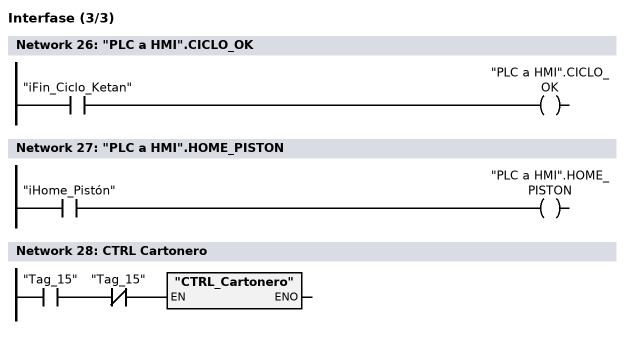
   RUNG wire#powerrail
      Contact( "iFin_Ciclo_Ketan" )
      Coil( "PLC a HMI".CICLO_OK )
   END_RUNG
   // the same network as SCL:
   "PLC a HMI".CICLO_OK := "iFin_Ciclo_Ketan";
END_REGION

REGION Network 27: "PLC a HMI".HOME_PISTON
   RUNG wire#powerrail
      Contact( "iHome_Pistón" )
      Coil( "PLC a HMI".HOME_PISTON )
   END_RUNG
   // the same network as SCL:
   "PLC a HMI".HOME_PISTON := "iHome_Pistón";
END_REGION

REGION Network 28: CTRL Cartonero
   RUNG wire#powerrail
      Contact( "Tag_15" )
      I_Contact( "Tag_15" )
      "CTRL_Cartonero"()
   END_RUNG
   // the same network as SCL:
   IF "Tag_15" AND NOT "Tag_15" THEN "CTRL_Cartonero"(); END_IF;
END_REGION
END_FUNCTION

FUNCTION "Conteo_AUTO" : Void   // FC26, STL
{ S7_Optimized_Access := 'FALSE' }
VERSION : 0.1
BEGIN

REGION Network 1: "Proceso CargaPallet".Capa_Actual
   // Con el fp del empujador adelante de todo, actualiza la "Capa_Actual" del grupo "CargaPalet"
         A     "flanco".piSnsEmpj_Ade_Par;
         JCN   NoCapa;
         L     "Proceso Empujador".Capa_Actual;
         T     "Proceso CargaPallet".Capa_Actual;
   NoCapa:NOP   0;
END_REGION

REGION Network 2
         L     "DB_Receta_Actual".Nro_Capas_Pallet;
         L     "Proceso Empujador".Capa_Actual;
         >I;
         =     #Habil_Inc;
         ==I;
         =     #Fin_Pallet;
         SET;
         A     #Habil_Inc;
         A     "flanco".piSnsEmpj_Ade_Par;
         JCN   noInc;
         L     "Proceso Empujador".Capa_Actual;
         INC   1;
         T     "Proceso Empujador".Capa_Actual;
   noInc:NOP   0;
         SET;
         A     #Fin_Pallet;
         A     "flanco".piSnsEmpj_Ade_Par;

         JCN   noFin;
         SET;
         S     "Última_Capa";
         L     1;
         T     "Proceso Empujador".Capa_Actual;
         L     "Proceso Empujador".Cant_Pallets;
         INC   1;
         T     "Proceso Empujador".Cant_Pallets;
   noFin:NOP   0;

         A     "flanco".nPALLET_NO_FUERA_ASCENSOR;
         JCN   noWRPall;
         L     "Proceso Empujador".Cant_Pallets;
         T     "Proceso CargaPallet".Cant_Pallets;
   noWRPall:NOP   0;


   //////////////////////////////
   //      O     "Ascensor_Zona_Superior"//
   //U     "flanco".nPALLET_NO_FUERA_ASCENSOR
   //     R     "Última_Capa"
END_REGION
END_FUNCTION

FUNCTION "Filtros_Señales" : Void   // FC27, LAD
{ S7_Optimized_Access := 'FALSE' }
VERSION : 0.1
BEGIN

REGION Network 1: Sensor Contador de embalaje 1
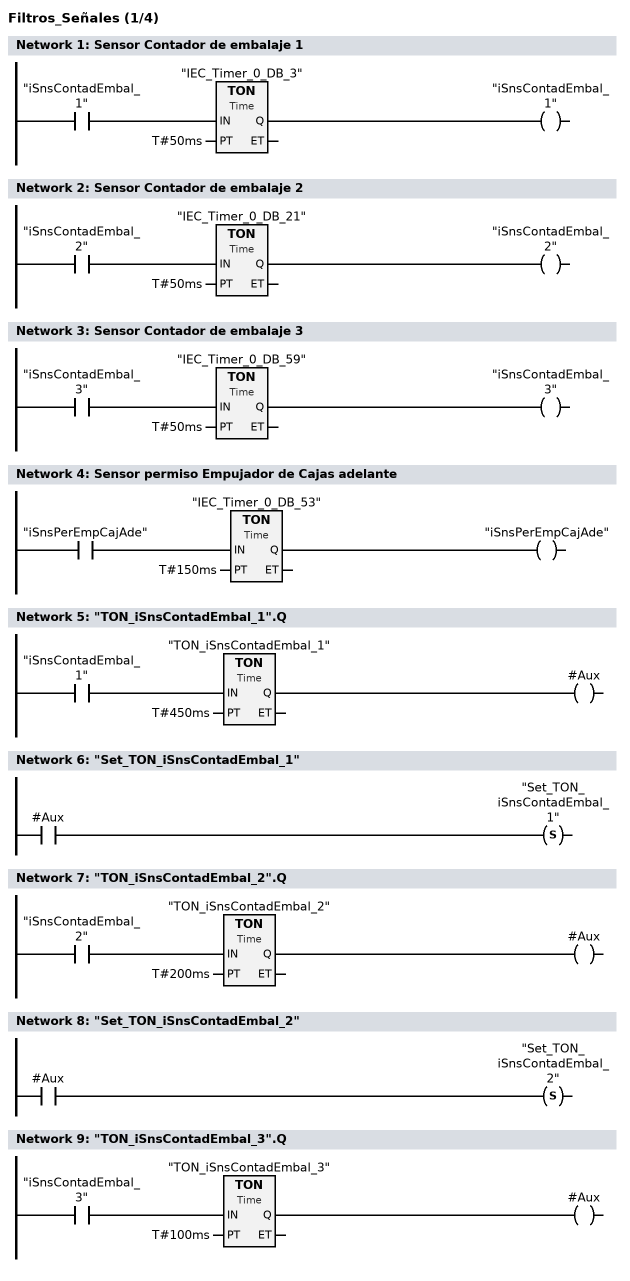
   "IEC_Timer_0_DB_3".TON(IN := "iSnsContadEmbal_1", PT := T#50ms);
   "iSnsContadEmbal_1" := "IEC_Timer_0_DB_3".Q;
END_REGION

REGION Network 2: Sensor Contador de embalaje 2
   "IEC_Timer_0_DB_21".TON(IN := "iSnsContadEmbal_2", PT := T#50ms);
   "iSnsContadEmbal_2" := "IEC_Timer_0_DB_21".Q;
END_REGION

REGION Network 3: Sensor Contador de embalaje 3
   "IEC_Timer_0_DB_59".TON(IN := "iSnsContadEmbal_3", PT := T#50ms);
   "iSnsContadEmbal_3" := "IEC_Timer_0_DB_59".Q;
END_REGION

REGION Network 4: Sensor permiso Empujador de Cajas adelante
   "IEC_Timer_0_DB_53".TON(IN := "iSnsPerEmpCajAde", PT := T#150ms);
   "iSnsPerEmpCajAde" := "IEC_Timer_0_DB_53".Q;
END_REGION

REGION Network 5: "TON_iSnsContadEmbal_1".Q
   "TON_iSnsContadEmbal_1".TON(IN := "iSnsContadEmbal_1", PT := T#450ms);
   #Aux := "TON_iSnsContadEmbal_1".Q;
END_REGION

REGION Network 6: "Set_TON_iSnsContadEmbal_1"
   RUNG wire#powerrail
      Contact( #Aux )
      S_Coil( "Set_TON_iSnsContadEmbal_1" )
   END_RUNG
   // the same network as SCL:
   IF #Aux THEN "Set_TON_iSnsContadEmbal_1" := TRUE; END_IF;
END_REGION

REGION Network 7: "TON_iSnsContadEmbal_2".Q
   "TON_iSnsContadEmbal_2".TON(IN := "iSnsContadEmbal_2", PT := T#200ms);
   #Aux := "TON_iSnsContadEmbal_2".Q;
END_REGION

REGION Network 8: "Set_TON_iSnsContadEmbal_2"
   RUNG wire#powerrail
      Contact( #Aux )
      S_Coil( "Set_TON_iSnsContadEmbal_2" )
   END_RUNG
   // the same network as SCL:
   IF #Aux THEN "Set_TON_iSnsContadEmbal_2" := TRUE; END_IF;
END_REGION

REGION Network 9: "TON_iSnsContadEmbal_3".Q
   "TON_iSnsContadEmbal_3".TON(IN := "iSnsContadEmbal_3", PT := T#100ms);
   #Aux := "TON_iSnsContadEmbal_3".Q;
END_REGION

REGION Network 10: "Set_TON_iSnsContadEmbal_3"
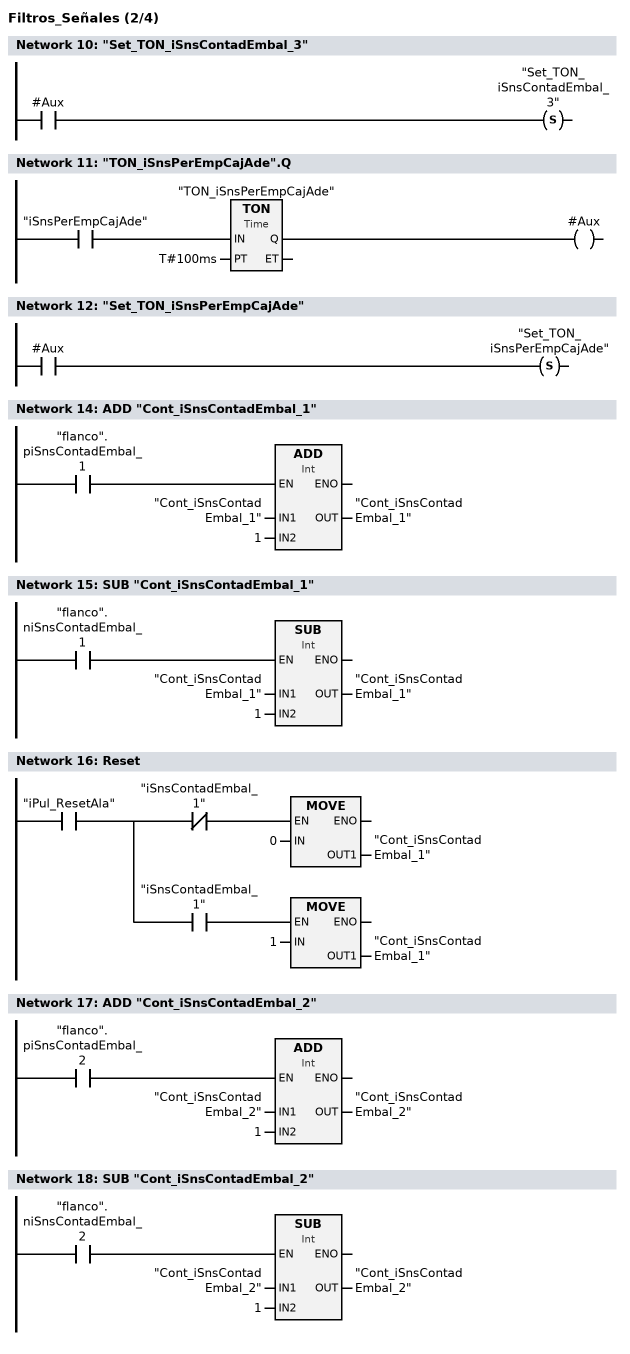
   RUNG wire#powerrail
      Contact( #Aux )
      S_Coil( "Set_TON_iSnsContadEmbal_3" )
   END_RUNG
   // the same network as SCL:
   IF #Aux THEN "Set_TON_iSnsContadEmbal_3" := TRUE; END_IF;
END_REGION

REGION Network 11: "TON_iSnsPerEmpCajAde".Q
   "TON_iSnsPerEmpCajAde".TON(IN := "iSnsPerEmpCajAde", PT := T#100ms);
   #Aux := "TON_iSnsPerEmpCajAde".Q;
END_REGION

REGION Network 12: "Set_TON_iSnsPerEmpCajAde"
   RUNG wire#powerrail
      Contact( #Aux )
      S_Coil( "Set_TON_iSnsPerEmpCajAde" )
   END_RUNG
   // the same network as SCL:
   IF #Aux THEN "Set_TON_iSnsPerEmpCajAde" := TRUE; END_IF;
END_REGION

REGION Network 13: ------------------------------------------ Control de flancos -------------------------------------------------
END_REGION

REGION Network 14: ADD "Cont_iSnsContadEmbal_1"
   RUNG wire#powerrail
      Contact( "flanco".piSnsContadEmbal_1 )
      { S7_Templates := "SrcType := Int"; S7_GenerateENO := "TRUE" } Add(in1 := "Cont_iSnsContadEmbal_1", in2 := 1, out => "Cont_iSnsContadEmbal_1")
   END_RUNG
   // the same network as SCL:
   IF "flanco".piSnsContadEmbal_1 THEN "Cont_iSnsContadEmbal_1" := "Cont_iSnsContadEmbal_1" + 1; END_IF;
END_REGION

REGION Network 15: SUB "Cont_iSnsContadEmbal_1"
   RUNG wire#powerrail
      Contact( "flanco".niSnsContadEmbal_1 )
      { S7_Templates := "SrcType := Int"; S7_GenerateENO := "TRUE" } Sub(in1 := "Cont_iSnsContadEmbal_1", in2 := 1, out => "Cont_iSnsContadEmbal_1")
   END_RUNG
   // the same network as SCL:
   IF "flanco".niSnsContadEmbal_1 THEN "Cont_iSnsContadEmbal_1" := "Cont_iSnsContadEmbal_1" - 1; END_IF;
END_REGION

REGION Network 16: Reset
   RUNG wire#powerrail
      Contact( "iPul_ResetAla" )
      wire#w1
      I_Contact( "iSnsContadEmbal_1" )
      { S7_GenerateENO := "TRUE" } Move(in := 0, out1 => "Cont_iSnsContadEmbal_1")
   END_RUNG
   RUNG wire#w1
      Contact( "iSnsContadEmbal_1" )
      { S7_GenerateENO := "TRUE" } Move(in := 1, out1 => "Cont_iSnsContadEmbal_1")
   END_RUNG
   // the same network as SCL:
   IF "iPul_ResetAla" AND NOT "iSnsContadEmbal_1" THEN "Cont_iSnsContadEmbal_1" := 0; END_IF;
   IF "iPul_ResetAla" AND "iSnsContadEmbal_1" THEN "Cont_iSnsContadEmbal_1" := 1; END_IF;
END_REGION

REGION Network 17: ADD "Cont_iSnsContadEmbal_2"
   RUNG wire#powerrail
      Contact( "flanco".piSnsContadEmbal_2 )
      { S7_Templates := "SrcType := Int"; S7_GenerateENO := "TRUE" } Add(in1 := "Cont_iSnsContadEmbal_2", in2 := 1, out => "Cont_iSnsContadEmbal_2")
   END_RUNG
   // the same network as SCL:
   IF "flanco".piSnsContadEmbal_2 THEN "Cont_iSnsContadEmbal_2" := "Cont_iSnsContadEmbal_2" + 1; END_IF;
END_REGION

REGION Network 18: SUB "Cont_iSnsContadEmbal_2"
   RUNG wire#powerrail
      Contact( "flanco".niSnsContadEmbal_2 )
      { S7_Templates := "SrcType := Int"; S7_GenerateENO := "TRUE" } Sub(in1 := "Cont_iSnsContadEmbal_2", in2 := 1, out => "Cont_iSnsContadEmbal_2")
   END_RUNG
   // the same network as SCL:
   IF "flanco".niSnsContadEmbal_2 THEN "Cont_iSnsContadEmbal_2" := "Cont_iSnsContadEmbal_2" - 1; END_IF;
END_REGION

REGION Network 19: Reset
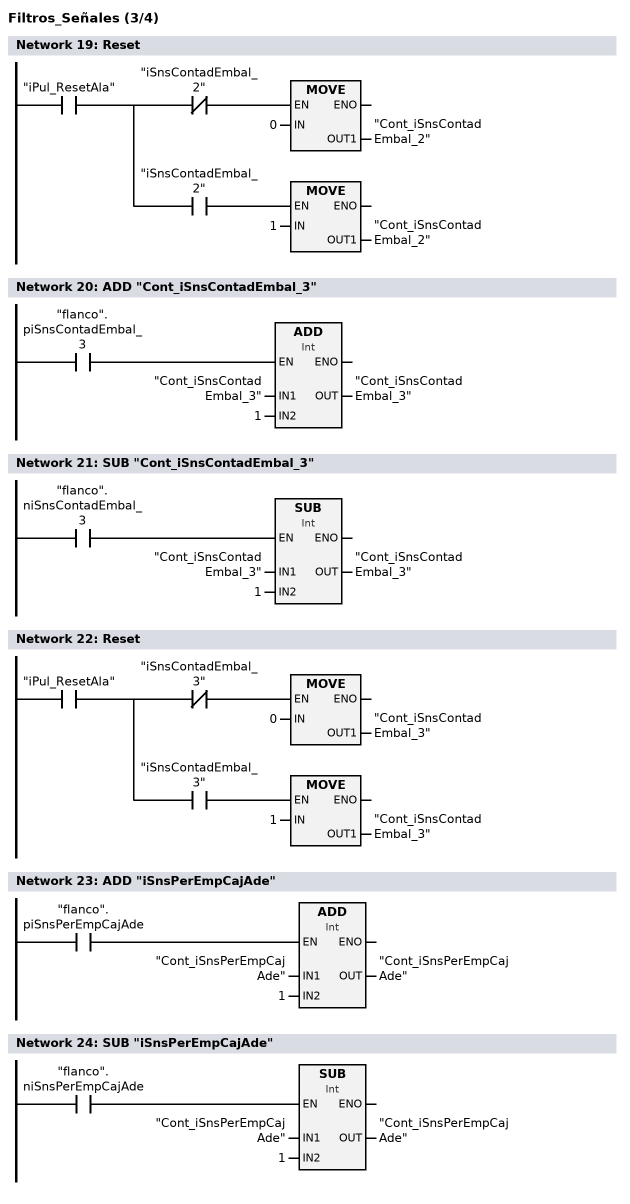
   RUNG wire#powerrail
      Contact( "iPul_ResetAla" )
      wire#w1
      I_Contact( "iSnsContadEmbal_2" )
      { S7_GenerateENO := "TRUE" } Move(in := 0, out1 => "Cont_iSnsContadEmbal_2")
   END_RUNG
   RUNG wire#w1
      Contact( "iSnsContadEmbal_2" )
      { S7_GenerateENO := "TRUE" } Move(in := 1, out1 => "Cont_iSnsContadEmbal_2")
   END_RUNG
   // the same network as SCL:
   IF "iPul_ResetAla" AND NOT "iSnsContadEmbal_2" THEN "Cont_iSnsContadEmbal_2" := 0; END_IF;
   IF "iPul_ResetAla" AND "iSnsContadEmbal_2" THEN "Cont_iSnsContadEmbal_2" := 1; END_IF;
END_REGION

REGION Network 20: ADD "Cont_iSnsContadEmbal_3"
   RUNG wire#powerrail
      Contact( "flanco".piSnsContadEmbal_3 )
      { S7_Templates := "SrcType := Int"; S7_GenerateENO := "TRUE" } Add(in1 := "Cont_iSnsContadEmbal_3", in2 := 1, out => "Cont_iSnsContadEmbal_3")
   END_RUNG
   // the same network as SCL:
   IF "flanco".piSnsContadEmbal_3 THEN "Cont_iSnsContadEmbal_3" := "Cont_iSnsContadEmbal_3" + 1; END_IF;
END_REGION

REGION Network 21: SUB "Cont_iSnsContadEmbal_3"
   RUNG wire#powerrail
      Contact( "flanco".niSnsContadEmbal_3 )
      { S7_Templates := "SrcType := Int"; S7_GenerateENO := "TRUE" } Sub(in1 := "Cont_iSnsContadEmbal_3", in2 := 1, out => "Cont_iSnsContadEmbal_3")
   END_RUNG
   // the same network as SCL:
   IF "flanco".niSnsContadEmbal_3 THEN "Cont_iSnsContadEmbal_3" := "Cont_iSnsContadEmbal_3" - 1; END_IF;
END_REGION

REGION Network 22: Reset
   RUNG wire#powerrail
      Contact( "iPul_ResetAla" )
      wire#w1
      I_Contact( "iSnsContadEmbal_3" )
      { S7_GenerateENO := "TRUE" } Move(in := 0, out1 => "Cont_iSnsContadEmbal_3")
   END_RUNG
   RUNG wire#w1
      Contact( "iSnsContadEmbal_3" )
      { S7_GenerateENO := "TRUE" } Move(in := 1, out1 => "Cont_iSnsContadEmbal_3")
   END_RUNG
   // the same network as SCL:
   IF "iPul_ResetAla" AND NOT "iSnsContadEmbal_3" THEN "Cont_iSnsContadEmbal_3" := 0; END_IF;
   IF "iPul_ResetAla" AND "iSnsContadEmbal_3" THEN "Cont_iSnsContadEmbal_3" := 1; END_IF;
END_REGION

REGION Network 23: ADD "iSnsPerEmpCajAde"
   RUNG wire#powerrail
      Contact( "flanco".piSnsPerEmpCajAde )
      { S7_Templates := "SrcType := Int"; S7_GenerateENO := "TRUE" } Add(in1 := "Cont_iSnsPerEmpCajAde", in2 := 1, out => "Cont_iSnsPerEmpCajAde")
   END_RUNG
   // the same network as SCL:
   IF "flanco".piSnsPerEmpCajAde THEN "Cont_iSnsPerEmpCajAde" := "Cont_iSnsPerEmpCajAde" + 1; END_IF;
END_REGION

REGION Network 24: SUB "iSnsPerEmpCajAde"
   RUNG wire#powerrail
      Contact( "flanco".niSnsPerEmpCajAde )
      { S7_Templates := "SrcType := Int"; S7_GenerateENO := "TRUE" } Sub(in1 := "Cont_iSnsPerEmpCajAde", in2 := 1, out => "Cont_iSnsPerEmpCajAde")
   END_RUNG
   // the same network as SCL:
   IF "flanco".niSnsPerEmpCajAde THEN "Cont_iSnsPerEmpCajAde" := "Cont_iSnsPerEmpCajAde" - 1; END_IF;
END_REGION

REGION Network 25: Reset
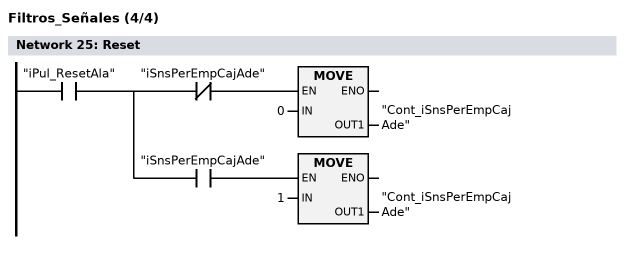
   RUNG wire#powerrail
      Contact( "iPul_ResetAla" )
      wire#w1
      I_Contact( "iSnsPerEmpCajAde" )
      { S7_GenerateENO := "TRUE" } Move(in := 0, out1 => "Cont_iSnsPerEmpCajAde")
   END_RUNG
   RUNG wire#w1
      Contact( "iSnsPerEmpCajAde" )
      { S7_GenerateENO := "TRUE" } Move(in := 1, out1 => "Cont_iSnsPerEmpCajAde")
   END_RUNG
   // the same network as SCL:
   IF "iPul_ResetAla" AND NOT "iSnsPerEmpCajAde" THEN "Cont_iSnsPerEmpCajAde" := 0; END_IF;
   IF "iPul_ResetAla" AND "iSnsPerEmpCajAde" THEN "Cont_iSnsPerEmpCajAde" := 1; END_IF;
END_REGION
END_FUNCTION

FUNCTION "CTRL_Cartonero" : Void   // FC29, LAD
{ S7_Optimized_Access := 'FALSE' }
VERSION : 0.1
BEGIN

REGION Network 1: Señal a Cartonero: 1= Tomar cartón
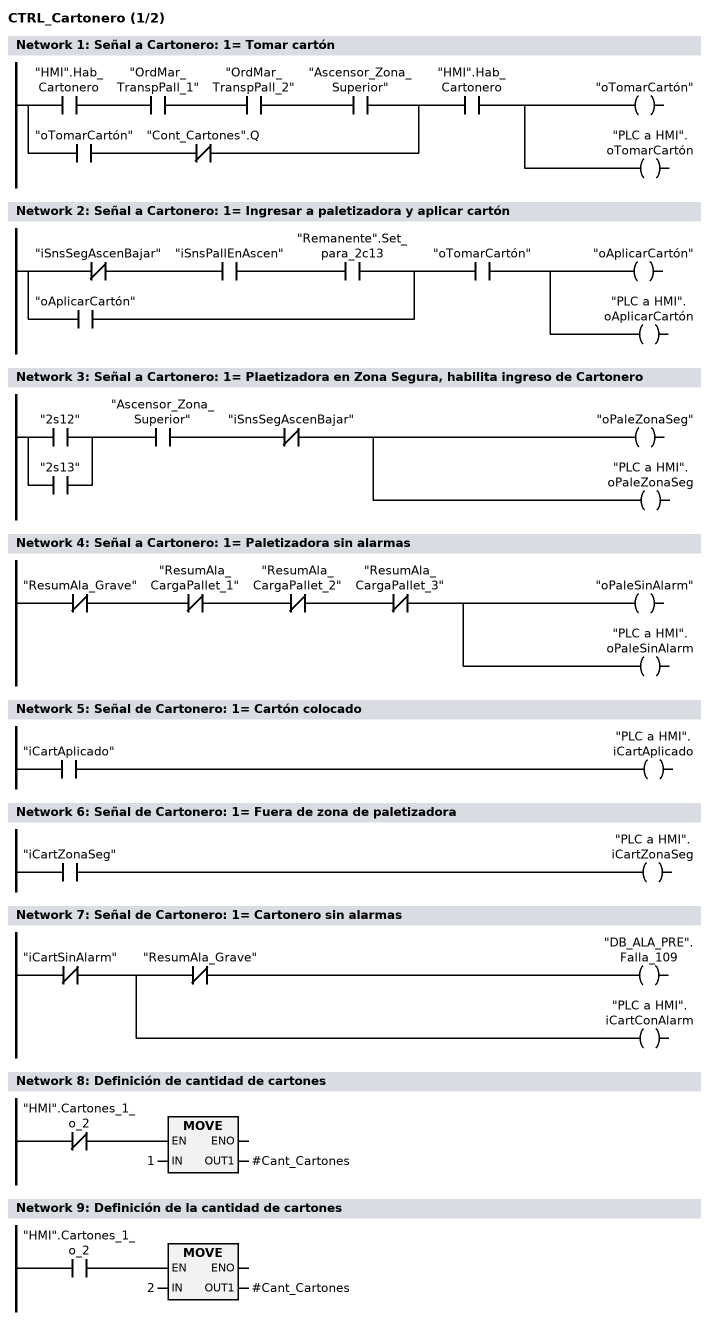
   RUNG wire#powerrail
      Contact( "HMI".Hab_Cartonero )
      Contact( "OrdMar_TranspPall_1" )
      Contact( "OrdMar_TranspPall_2" )
      Contact( "Ascensor_Zona_Superior" )
      wire#w1
      Contact( "HMI".Hab_Cartonero )
      wire#w2
      Coil( "oTomarCartón" )
   END_RUNG
   RUNG wire#powerrail
      Contact( "oTomarCartón" )
      I_Contact( "Cont_Cartones".Q )
   END_RUNG wire#w1
   RUNG wire#w2
      Coil( "PLC a HMI".oTomarCartón )
   END_RUNG
   // the same network as SCL:
   "oTomarCartón" := (("HMI".Hab_Cartonero AND "OrdMar_TranspPall_1" AND "OrdMar_TranspPall_2" AND "Ascensor_Zona_Superior") OR ("oTomarCartón" AND NOT "Cont_Cartones".Q)) AND "HMI".Hab_Cartonero;
   "PLC a HMI".oTomarCartón := "oTomarCartón";
END_REGION

REGION Network 2: Señal a Cartonero: 1= Ingresar a paletizadora y aplicar cartón
   RUNG wire#powerrail
      I_Contact( "iSnsSegAscenBajar" )
      Contact( "iSnsPallEnAscen" )
      Contact( "Remanente".Set_para_2c13 )
      wire#w1
      Contact( "oTomarCartón" )
      wire#w2
      Coil( "oAplicarCartón" )
   END_RUNG
   RUNG wire#powerrail
      Contact( "oAplicarCartón" )
   END_RUNG wire#w1
   RUNG wire#w2
      Coil( "PLC a HMI".oAplicarCartón )
   END_RUNG
   // the same network as SCL:
   "oAplicarCartón" := ((NOT "iSnsSegAscenBajar" AND "iSnsPallEnAscen" AND "Remanente".Set_para_2c13) OR "oAplicarCartón") AND "oTomarCartón";
   "PLC a HMI".oAplicarCartón := "oAplicarCartón";
END_REGION

REGION Network 3: Señal a Cartonero: 1= Plaetizadora en Zona Segura, habilita ingreso de Cartonero
   RUNG wire#powerrail
      Contact( "2s12" )
      wire#w1
      Contact( "Ascensor_Zona_Superior" )
      I_Contact( "iSnsSegAscenBajar" )
      wire#w2
      Coil( "oPaleZonaSeg" )
   END_RUNG
   RUNG wire#powerrail
      Contact( "2s13" )
   END_RUNG wire#w1
   RUNG wire#w2
      Coil( "PLC a HMI".oPaleZonaSeg )
   END_RUNG
   // the same network as SCL:
   "oPaleZonaSeg" := ("2s12" OR "2s13") AND "Ascensor_Zona_Superior" AND NOT "iSnsSegAscenBajar";
   "PLC a HMI".oPaleZonaSeg := "oPaleZonaSeg";
END_REGION

REGION Network 4: Señal a Cartonero: 1= Paletizadora sin alarmas
   RUNG wire#powerrail
      I_Contact( "ResumAla_Grave" )
      I_Contact( "ResumAla_CargaPallet_1" )
      I_Contact( "ResumAla_CargaPallet_2" )
      I_Contact( "ResumAla_CargaPallet_3" )
      wire#w1
      Coil( "oPaleSinAlarm" )
   END_RUNG
   RUNG wire#w1
      Coil( "PLC a HMI".oPaleSinAlarm )
   END_RUNG
   // the same network as SCL:
   "oPaleSinAlarm" := NOT "ResumAla_Grave" AND NOT "ResumAla_CargaPallet_1" AND NOT "ResumAla_CargaPallet_2" AND NOT "ResumAla_CargaPallet_3";
   "PLC a HMI".oPaleSinAlarm := "oPaleSinAlarm";
END_REGION

REGION Network 5: Señal de Cartonero: 1= Cartón colocado
   RUNG wire#powerrail
      Contact( "iCartAplicado" )
      Coil( "PLC a HMI".iCartAplicado )
   END_RUNG
   // the same network as SCL:
   "PLC a HMI".iCartAplicado := "iCartAplicado";
END_REGION

REGION Network 6: Señal de Cartonero: 1= Fuera de zona de paletizadora
   RUNG wire#powerrail
      Contact( "iCartZonaSeg" )
      Coil( "PLC a HMI".iCartZonaSeg )
   END_RUNG
   // the same network as SCL:
   "PLC a HMI".iCartZonaSeg := "iCartZonaSeg";
END_REGION

REGION Network 7: Señal de Cartonero: 1= Cartonero sin alarmas
   RUNG wire#powerrail
      I_Contact( "iCartSinAlarm" )
      wire#w1
      I_Contact( "ResumAla_Grave" )
      Coil( "DB_ALA_PRE".Falla_109 )
   END_RUNG
   RUNG wire#w1
      Coil( "PLC a HMI".iCartConAlarm )
   END_RUNG
   // the same network as SCL:
   "DB_ALA_PRE".Falla_109 := NOT "iCartSinAlarm" AND NOT "ResumAla_Grave";
   "PLC a HMI".iCartConAlarm := NOT "iCartSinAlarm";
END_REGION

REGION Network 8: Definición de cantidad de cartones
   RUNG wire#powerrail
      I_Contact( "HMI".Cartones_1_o_2 )
      { S7_GenerateENO := "TRUE" } Move(in := 1, out1 => #Cant_Cartones)
   END_RUNG
   // the same network as SCL:
   IF NOT "HMI".Cartones_1_o_2 THEN #Cant_Cartones := 1; END_IF;
END_REGION

REGION Network 9: Definición de la cantidad de cartones
   RUNG wire#powerrail
      Contact( "HMI".Cartones_1_o_2 )
      { S7_GenerateENO := "TRUE" } Move(in := 2, out1 => #Cant_Cartones)
   END_RUNG
   // the same network as SCL:
   IF "HMI".Cartones_1_o_2 THEN #Cant_Cartones := 2; END_IF;
END_REGION

REGION Network 10: Contador cartones
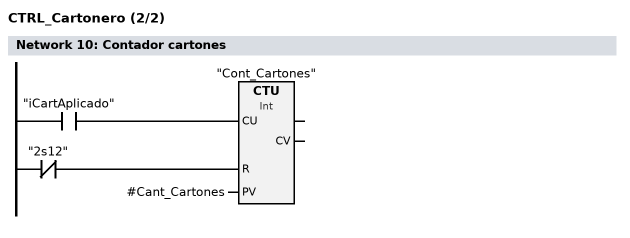
   "Cont_Cartones".CTU(CU := "iCartAplicado", R := NOT "2s12", PV := #Cant_Cartones);
END_REGION
END_FUNCTION

FUNCTION "ReparaRecetas_Pistón" : Void   // FC30, LAD
{ S7_Optimized_Access := 'FALSE' }
VERSION : 0.1
BEGIN

REGION Network 1: Repara receta 1
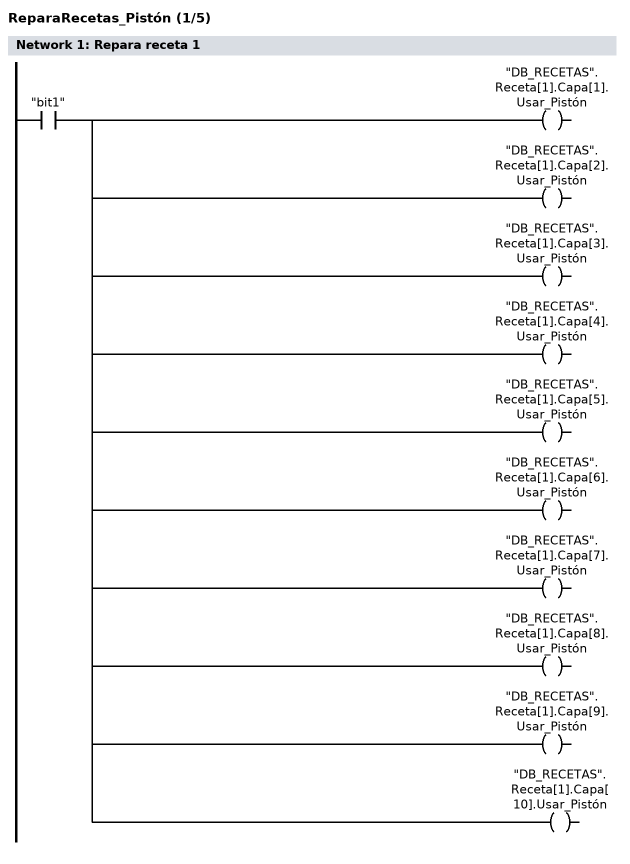
   RUNG wire#powerrail
      Contact( "bit1" )
      wire#w1
      Coil( "DB_RECETAS".Receta[1].Capa[1].Usar_Pistón )
   END_RUNG
   RUNG wire#w1
      Coil( "DB_RECETAS".Receta[1].Capa[2].Usar_Pistón )
   END_RUNG
   RUNG wire#w1
      Coil( "DB_RECETAS".Receta[1].Capa[3].Usar_Pistón )
   END_RUNG
   RUNG wire#w1
      Coil( "DB_RECETAS".Receta[1].Capa[4].Usar_Pistón )
   END_RUNG
   RUNG wire#w1
      Coil( "DB_RECETAS".Receta[1].Capa[5].Usar_Pistón )
   END_RUNG
   RUNG wire#w1
      Coil( "DB_RECETAS".Receta[1].Capa[6].Usar_Pistón )
   END_RUNG
   RUNG wire#w1
      Coil( "DB_RECETAS".Receta[1].Capa[7].Usar_Pistón )
   END_RUNG
   RUNG wire#w1
      Coil( "DB_RECETAS".Receta[1].Capa[8].Usar_Pistón )
   END_RUNG
   RUNG wire#w1
      Coil( "DB_RECETAS".Receta[1].Capa[9].Usar_Pistón )
   END_RUNG
   RUNG wire#w1
      Coil( "DB_RECETAS".Receta[1].Capa[10].Usar_Pistón )
   END_RUNG
   // the same network as SCL:
   "DB_RECETAS".Receta[1].Capa[1].Usar_Pistón := "bit1";
   "DB_RECETAS".Receta[1].Capa[2].Usar_Pistón := "bit1";
   "DB_RECETAS".Receta[1].Capa[3].Usar_Pistón := "bit1";
   "DB_RECETAS".Receta[1].Capa[4].Usar_Pistón := "bit1";
   "DB_RECETAS".Receta[1].Capa[5].Usar_Pistón := "bit1";
   "DB_RECETAS".Receta[1].Capa[6].Usar_Pistón := "bit1";
   "DB_RECETAS".Receta[1].Capa[7].Usar_Pistón := "bit1";
   "DB_RECETAS".Receta[1].Capa[8].Usar_Pistón := "bit1";
   "DB_RECETAS".Receta[1].Capa[9].Usar_Pistón := "bit1";
   "DB_RECETAS".Receta[1].Capa[10].Usar_Pistón := "bit1";
END_REGION

REGION Network 2: Repara receta 3
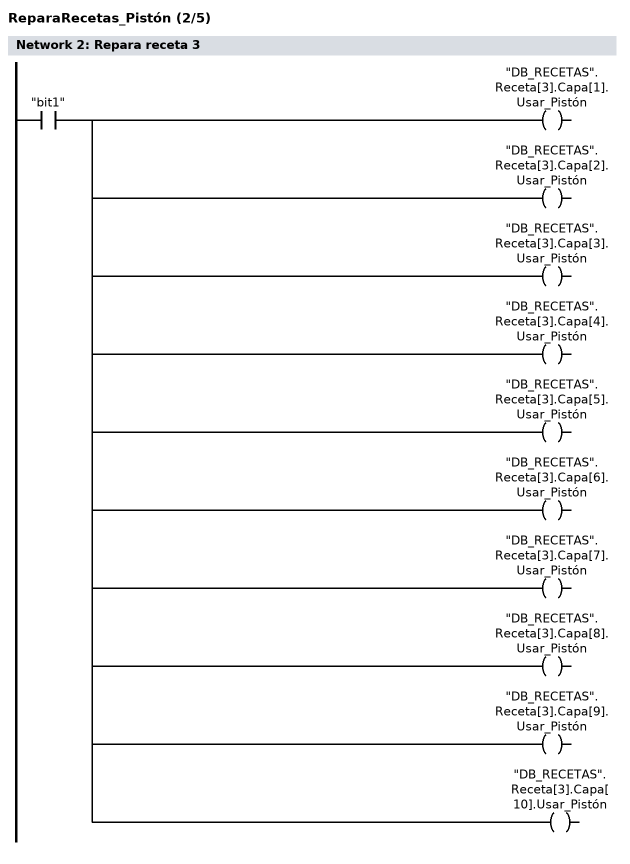
   RUNG wire#powerrail
      Contact( "bit1" )
      wire#w1
      Coil( "DB_RECETAS".Receta[3].Capa[1].Usar_Pistón )
   END_RUNG
   RUNG wire#w1
      Coil( "DB_RECETAS".Receta[3].Capa[2].Usar_Pistón )
   END_RUNG
   RUNG wire#w1
      Coil( "DB_RECETAS".Receta[3].Capa[3].Usar_Pistón )
   END_RUNG
   RUNG wire#w1
      Coil( "DB_RECETAS".Receta[3].Capa[4].Usar_Pistón )
   END_RUNG
   RUNG wire#w1
      Coil( "DB_RECETAS".Receta[3].Capa[5].Usar_Pistón )
   END_RUNG
   RUNG wire#w1
      Coil( "DB_RECETAS".Receta[3].Capa[6].Usar_Pistón )
   END_RUNG
   RUNG wire#w1
      Coil( "DB_RECETAS".Receta[3].Capa[7].Usar_Pistón )
   END_RUNG
   RUNG wire#w1
      Coil( "DB_RECETAS".Receta[3].Capa[8].Usar_Pistón )
   END_RUNG
   RUNG wire#w1
      Coil( "DB_RECETAS".Receta[3].Capa[9].Usar_Pistón )
   END_RUNG
   RUNG wire#w1
      Coil( "DB_RECETAS".Receta[3].Capa[10].Usar_Pistón )
   END_RUNG
   // the same network as SCL:
   "DB_RECETAS".Receta[3].Capa[1].Usar_Pistón := "bit1";
   "DB_RECETAS".Receta[3].Capa[2].Usar_Pistón := "bit1";
   "DB_RECETAS".Receta[3].Capa[3].Usar_Pistón := "bit1";
   "DB_RECETAS".Receta[3].Capa[4].Usar_Pistón := "bit1";
   "DB_RECETAS".Receta[3].Capa[5].Usar_Pistón := "bit1";
   "DB_RECETAS".Receta[3].Capa[6].Usar_Pistón := "bit1";
   "DB_RECETAS".Receta[3].Capa[7].Usar_Pistón := "bit1";
   "DB_RECETAS".Receta[3].Capa[8].Usar_Pistón := "bit1";
   "DB_RECETAS".Receta[3].Capa[9].Usar_Pistón := "bit1";
   "DB_RECETAS".Receta[3].Capa[10].Usar_Pistón := "bit1";
END_REGION

REGION Network 3: Repara receta 4
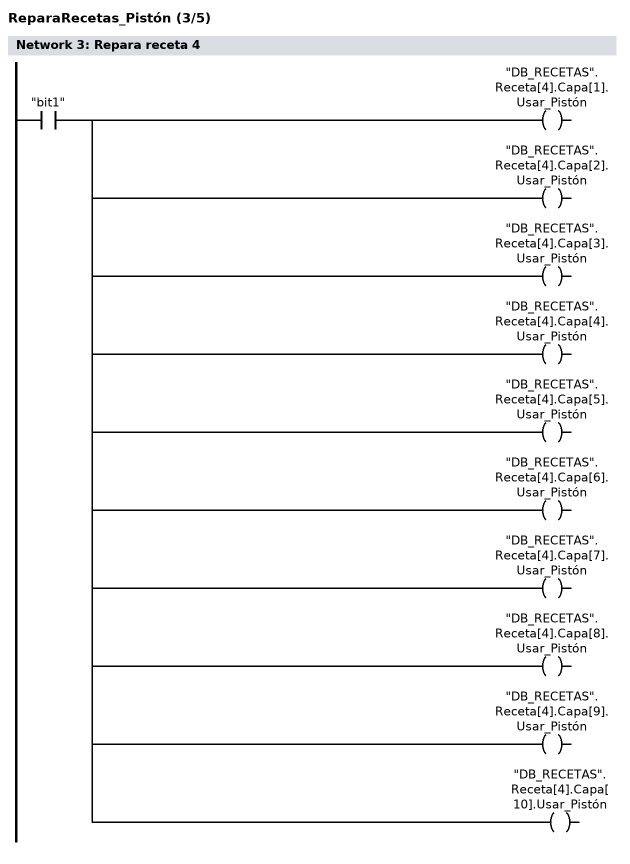
   RUNG wire#powerrail
      Contact( "bit1" )
      wire#w1
      Coil( "DB_RECETAS".Receta[4].Capa[1].Usar_Pistón )
   END_RUNG
   RUNG wire#w1
      Coil( "DB_RECETAS".Receta[4].Capa[2].Usar_Pistón )
   END_RUNG
   RUNG wire#w1
      Coil( "DB_RECETAS".Receta[4].Capa[3].Usar_Pistón )
   END_RUNG
   RUNG wire#w1
      Coil( "DB_RECETAS".Receta[4].Capa[4].Usar_Pistón )
   END_RUNG
   RUNG wire#w1
      Coil( "DB_RECETAS".Receta[4].Capa[5].Usar_Pistón )
   END_RUNG
   RUNG wire#w1
      Coil( "DB_RECETAS".Receta[4].Capa[6].Usar_Pistón )
   END_RUNG
   RUNG wire#w1
      Coil( "DB_RECETAS".Receta[4].Capa[7].Usar_Pistón )
   END_RUNG
   RUNG wire#w1
      Coil( "DB_RECETAS".Receta[4].Capa[8].Usar_Pistón )
   END_RUNG
   RUNG wire#w1
      Coil( "DB_RECETAS".Receta[4].Capa[9].Usar_Pistón )
   END_RUNG
   RUNG wire#w1
      Coil( "DB_RECETAS".Receta[4].Capa[10].Usar_Pistón )
   END_RUNG
   // the same network as SCL:
   "DB_RECETAS".Receta[4].Capa[1].Usar_Pistón := "bit1";
   "DB_RECETAS".Receta[4].Capa[2].Usar_Pistón := "bit1";
   "DB_RECETAS".Receta[4].Capa[3].Usar_Pistón := "bit1";
   "DB_RECETAS".Receta[4].Capa[4].Usar_Pistón := "bit1";
   "DB_RECETAS".Receta[4].Capa[5].Usar_Pistón := "bit1";
   "DB_RECETAS".Receta[4].Capa[6].Usar_Pistón := "bit1";
   "DB_RECETAS".Receta[4].Capa[7].Usar_Pistón := "bit1";
   "DB_RECETAS".Receta[4].Capa[8].Usar_Pistón := "bit1";
   "DB_RECETAS".Receta[4].Capa[9].Usar_Pistón := "bit1";
   "DB_RECETAS".Receta[4].Capa[10].Usar_Pistón := "bit1";
END_REGION

REGION Network 4: Repara receta 5
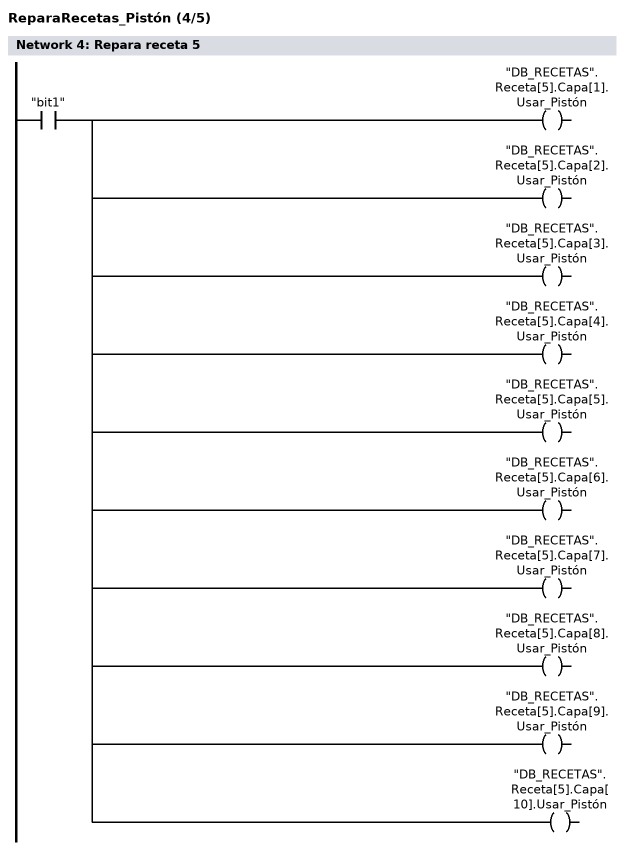
   RUNG wire#powerrail
      Contact( "bit1" )
      wire#w1
      Coil( "DB_RECETAS".Receta[5].Capa[1].Usar_Pistón )
   END_RUNG
   RUNG wire#w1
      Coil( "DB_RECETAS".Receta[5].Capa[2].Usar_Pistón )
   END_RUNG
   RUNG wire#w1
      Coil( "DB_RECETAS".Receta[5].Capa[3].Usar_Pistón )
   END_RUNG
   RUNG wire#w1
      Coil( "DB_RECETAS".Receta[5].Capa[4].Usar_Pistón )
   END_RUNG
   RUNG wire#w1
      Coil( "DB_RECETAS".Receta[5].Capa[5].Usar_Pistón )
   END_RUNG
   RUNG wire#w1
      Coil( "DB_RECETAS".Receta[5].Capa[6].Usar_Pistón )
   END_RUNG
   RUNG wire#w1
      Coil( "DB_RECETAS".Receta[5].Capa[7].Usar_Pistón )
   END_RUNG
   RUNG wire#w1
      Coil( "DB_RECETAS".Receta[5].Capa[8].Usar_Pistón )
   END_RUNG
   RUNG wire#w1
      Coil( "DB_RECETAS".Receta[5].Capa[9].Usar_Pistón )
   END_RUNG
   RUNG wire#w1
      Coil( "DB_RECETAS".Receta[5].Capa[10].Usar_Pistón )
   END_RUNG
   // the same network as SCL:
   "DB_RECETAS".Receta[5].Capa[1].Usar_Pistón := "bit1";
   "DB_RECETAS".Receta[5].Capa[2].Usar_Pistón := "bit1";
   "DB_RECETAS".Receta[5].Capa[3].Usar_Pistón := "bit1";
   "DB_RECETAS".Receta[5].Capa[4].Usar_Pistón := "bit1";
   "DB_RECETAS".Receta[5].Capa[5].Usar_Pistón := "bit1";
   "DB_RECETAS".Receta[5].Capa[6].Usar_Pistón := "bit1";
   "DB_RECETAS".Receta[5].Capa[7].Usar_Pistón := "bit1";
   "DB_RECETAS".Receta[5].Capa[8].Usar_Pistón := "bit1";
   "DB_RECETAS".Receta[5].Capa[9].Usar_Pistón := "bit1";
   "DB_RECETAS".Receta[5].Capa[10].Usar_Pistón := "bit1";
END_REGION

REGION Network 5: Repara receta 6
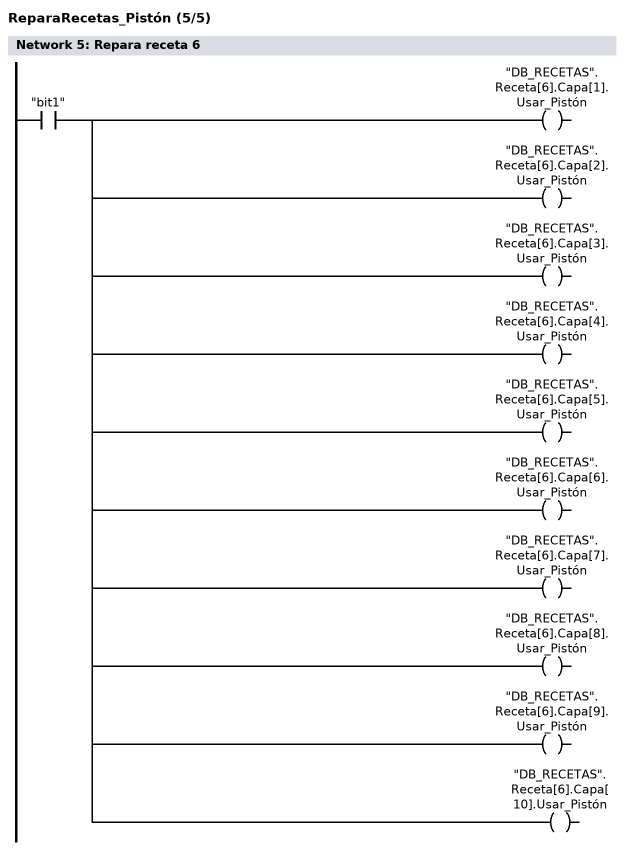
   RUNG wire#powerrail
      Contact( "bit1" )
      wire#w1
      Coil( "DB_RECETAS".Receta[6].Capa[1].Usar_Pistón )
   END_RUNG
   RUNG wire#w1
      Coil( "DB_RECETAS".Receta[6].Capa[2].Usar_Pistón )
   END_RUNG
   RUNG wire#w1
      Coil( "DB_RECETAS".Receta[6].Capa[3].Usar_Pistón )
   END_RUNG
   RUNG wire#w1
      Coil( "DB_RECETAS".Receta[6].Capa[4].Usar_Pistón )
   END_RUNG
   RUNG wire#w1
      Coil( "DB_RECETAS".Receta[6].Capa[5].Usar_Pistón )
   END_RUNG
   RUNG wire#w1
      Coil( "DB_RECETAS".Receta[6].Capa[6].Usar_Pistón )
   END_RUNG
   RUNG wire#w1
      Coil( "DB_RECETAS".Receta[6].Capa[7].Usar_Pistón )
   END_RUNG
   RUNG wire#w1
      Coil( "DB_RECETAS".Receta[6].Capa[8].Usar_Pistón )
   END_RUNG
   RUNG wire#w1
      Coil( "DB_RECETAS".Receta[6].Capa[9].Usar_Pistón )
   END_RUNG
   RUNG wire#w1
      Coil( "DB_RECETAS".Receta[6].Capa[10].Usar_Pistón )
   END_RUNG
   // the same network as SCL:
   "DB_RECETAS".Receta[6].Capa[1].Usar_Pistón := "bit1";
   "DB_RECETAS".Receta[6].Capa[2].Usar_Pistón := "bit1";
   "DB_RECETAS".Receta[6].Capa[3].Usar_Pistón := "bit1";
   "DB_RECETAS".Receta[6].Capa[4].Usar_Pistón := "bit1";
   "DB_RECETAS".Receta[6].Capa[5].Usar_Pistón := "bit1";
   "DB_RECETAS".Receta[6].Capa[6].Usar_Pistón := "bit1";
   "DB_RECETAS".Receta[6].Capa[7].Usar_Pistón := "bit1";
   "DB_RECETAS".Receta[6].Capa[8].Usar_Pistón := "bit1";
   "DB_RECETAS".Receta[6].Capa[9].Usar_Pistón := "bit1";
   "DB_RECETAS".Receta[6].Capa[10].Usar_Pistón := "bit1";
END_REGION
END_FUNCTION

ORGANIZATION_BLOCK "Main"   // OB1, LAD
TITLE = "Main Program Sweep (Cycle)"
{ S7_Optimized_Access := 'FALSE' }
VERSION : 0.1
BEGIN

REGION Network 1: Leer fecha y hora plc
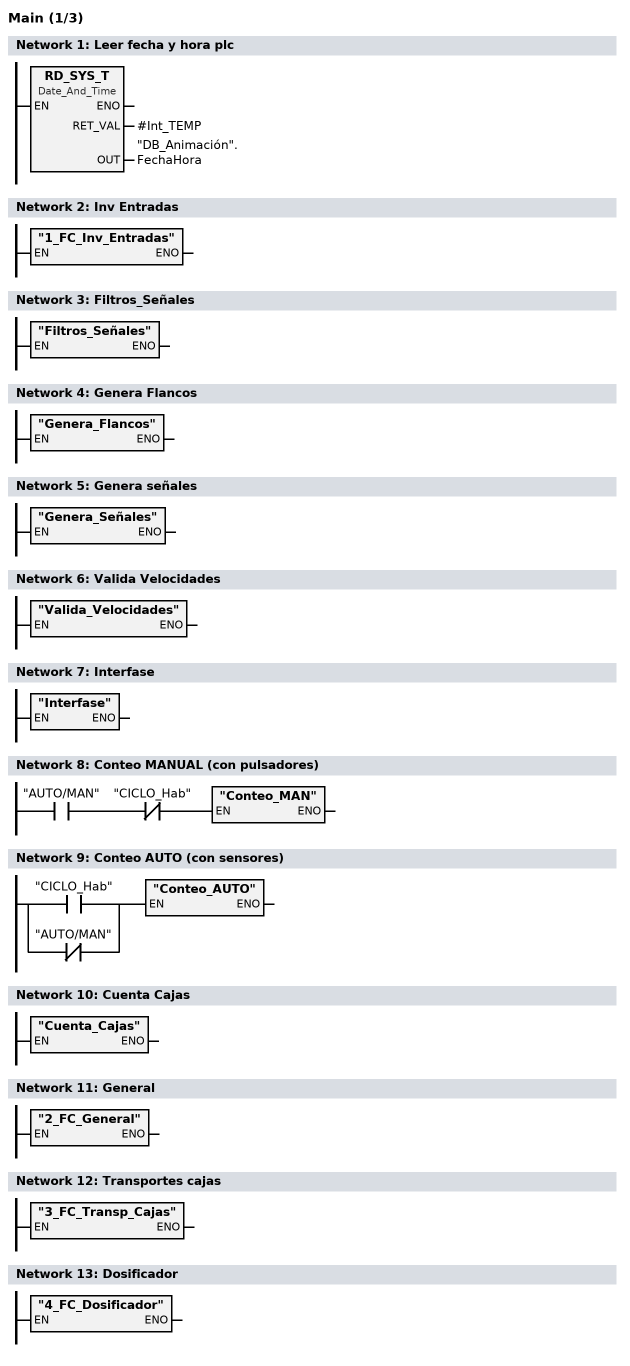
   #Int_TEMP := RD_SYS_T(out => "DB_Animación".FechaHora);
END_REGION

REGION Network 2: Inv Entradas
   RUNG wire#powerrail
      "1_FC_Inv_Entradas"()
   END_RUNG
   // the same network as SCL:
   "1_FC_Inv_Entradas"();
END_REGION

REGION Network 3: Filtros_Señales
   RUNG wire#powerrail
      "Filtros_Señales"()
   END_RUNG
   // the same network as SCL:
   "Filtros_Señales"();
END_REGION

REGION Network 4: Genera Flancos
   RUNG wire#powerrail
      "Genera_Flancos"()
   END_RUNG
   // the same network as SCL:
   "Genera_Flancos"();
END_REGION

REGION Network 5: Genera señales
   RUNG wire#powerrail
      "Genera_Señales"()
   END_RUNG
   // the same network as SCL:
   "Genera_Señales"();
END_REGION

REGION Network 6: Valida Velocidades
   RUNG wire#powerrail
      "Valida_Velocidades"()
   END_RUNG
   // the same network as SCL:
   "Valida_Velocidades"();
END_REGION

REGION Network 7: Interfase
   RUNG wire#powerrail
      "Interfase"()
   END_RUNG
   // the same network as SCL:
   "Interfase"();
END_REGION

REGION Network 8: Conteo MANUAL (con pulsadores)
   RUNG wire#powerrail
      Contact( "AUTO/MAN" )
      I_Contact( "CICLO_Hab" )
      "Conteo_MAN"()
   END_RUNG
   // the same network as SCL:
   IF "AUTO/MAN" AND NOT "CICLO_Hab" THEN "Conteo_MAN"(); END_IF;
END_REGION

REGION Network 9: Conteo AUTO (con sensores)
   RUNG wire#powerrail
      Contact( "CICLO_Hab" )
      wire#w1
      "Conteo_AUTO"()
   END_RUNG
   RUNG wire#powerrail
      I_Contact( "AUTO/MAN" )
   END_RUNG wire#w1
   // the same network as SCL:
   IF "CICLO_Hab" OR NOT "AUTO/MAN" THEN "Conteo_AUTO"(); END_IF;
END_REGION

REGION Network 10: Cuenta Cajas
   RUNG wire#powerrail
      "Cuenta_Cajas"()
   END_RUNG
   // the same network as SCL:
   "Cuenta_Cajas"();
END_REGION

REGION Network 11: General
   RUNG wire#powerrail
      "2_FC_General"()
   END_RUNG
   // the same network as SCL:
   "2_FC_General"();
END_REGION

REGION Network 12: Transportes cajas
   RUNG wire#powerrail
      "3_FC_Transp_Cajas"()
   END_RUNG
   // the same network as SCL:
   "3_FC_Transp_Cajas"();
END_REGION

REGION Network 13: Dosificador
   RUNG wire#powerrail
      "4_FC_Dosificador"()
   END_RUNG
   // the same network as SCL:
   "4_FC_Dosificador"();
END_REGION

REGION Network 14: ELEMENTO HH
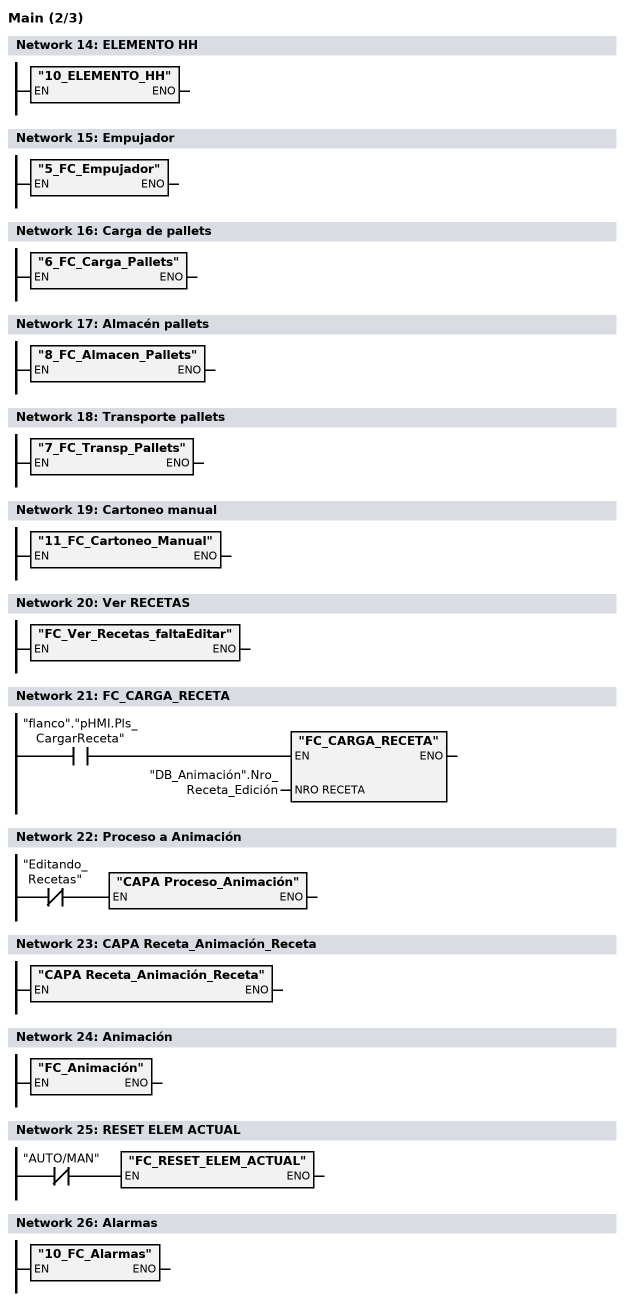
   RUNG wire#powerrail
      "10_ELEMENTO_HH"()
   END_RUNG
   // the same network as SCL:
   "10_ELEMENTO_HH"();
END_REGION

REGION Network 15: Empujador
   RUNG wire#powerrail
      "5_FC_Empujador"()
   END_RUNG
   // the same network as SCL:
   "5_FC_Empujador"();
END_REGION

REGION Network 16: Carga de pallets
   RUNG wire#powerrail
      "6_FC_Carga_Pallets"()
   END_RUNG
   // the same network as SCL:
   "6_FC_Carga_Pallets"();
END_REGION

REGION Network 17: Almacén pallets
   RUNG wire#powerrail
      "8_FC_Almacen_Pallets"()
   END_RUNG
   // the same network as SCL:
   "8_FC_Almacen_Pallets"();
END_REGION

REGION Network 18: Transporte pallets
   RUNG wire#powerrail
      "7_FC_Transp_Pallets"()
   END_RUNG
   // the same network as SCL:
   "7_FC_Transp_Pallets"();
END_REGION

REGION Network 19: Cartoneo manual
   RUNG wire#powerrail
      "11_FC_Cartoneo_Manual"()
   END_RUNG
   // the same network as SCL:
   "11_FC_Cartoneo_Manual"();
END_REGION

REGION Network 20: Ver RECETAS
   RUNG wire#powerrail
      "FC_Ver_Recetas_faltaEditar"()
   END_RUNG
   // the same network as SCL:
   "FC_Ver_Recetas_faltaEditar"();
END_REGION
